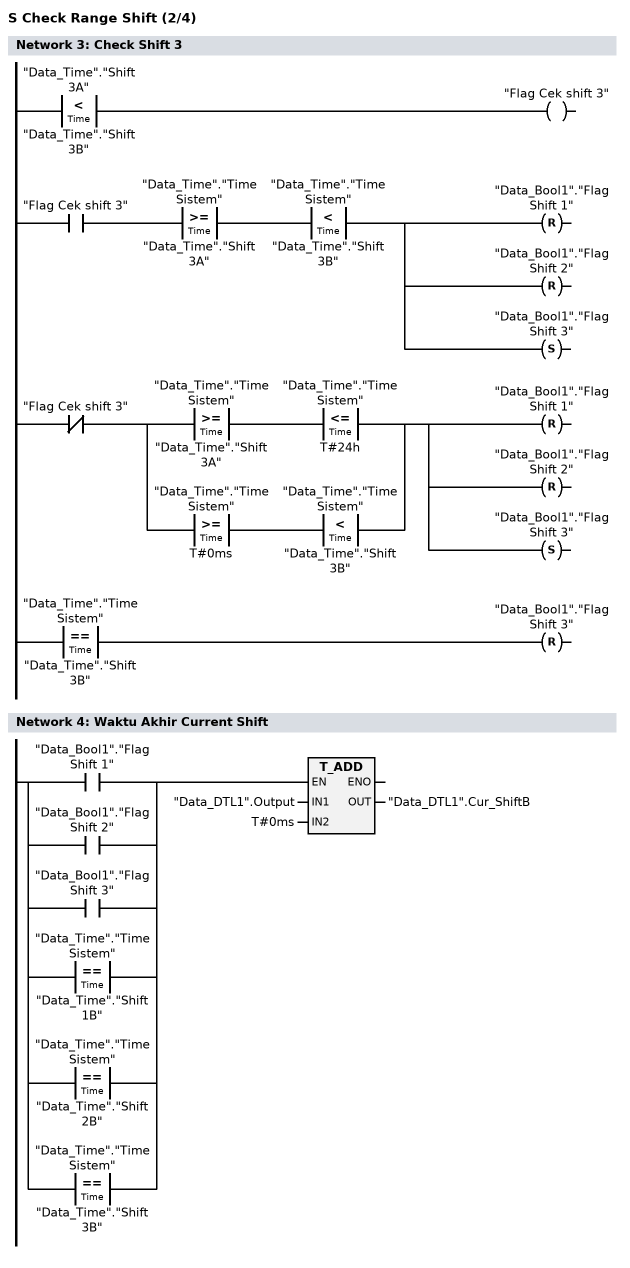
   RUNG wire#powerrail
      { S7_Templates := "SrcType := Time" } LT_Contact(in1 := "Data_Time"."Shift 3A", in2 := "Data_Time"."Shift 3B")
      Coil( "Flag Cek shift 3" )
   END_RUNG
   RUNG wire#powerrail
      Contact( "Flag Cek shift 3" )
      { S7_Templates := "SrcType := Time" } GE_Contact(in1 := "Data_Time"."Time Sistem", in2 := "Data_Time"."Shift 3A")
      { S7_Templates := "SrcType := Time" } LT_Contact(in1 := "Data_Time"."Time Sistem", in2 := "Data_Time"."Shift 3B")
      wire#w1
      R_Coil( "Data_Bool1"."Flag Shift 1" )
   END_RUNG
   RUNG wire#w1
      R_Coil( "Data_Bool1"."Flag Shift 2" )
   END_RUNG
   RUNG wire#w1
      S_Coil( "Data_Bool1"."Flag Shift 3" )
   END_RUNG
   RUNG wire#powerrail
      I_Contact( "Flag Cek shift 3" )
      wire#w2
      { S7_Templates := "SrcType := Time" } GE_Contact(in1 := "Data_Time"."Time Sistem", in2 := "Data_Time"."Shift 3A")
      { S7_Templates := "SrcType := Time" } LE_Contact(in1 := "Data_Time"."Time Sistem", in2 := T#24h)
      wire#w3
      R_Coil( "Data_Bool1"."Flag Shift 1" )
   END_RUNG
   RUNG wire#w2
      { S7_Templates := "SrcType := Time" } GE_Contact(in1 := "Data_Time"."Time Sistem", in2 := T#0ms)
      { S7_Templates := "SrcType := Time" } LT_Contact(in1 := "Data_Time"."Time Sistem", in2 := "Data_Time"."Shift 3B")
   END_RUNG wire#w3
   RUNG wire#w3
      R_Coil( "Data_Bool1"."Flag Shift 2" )
   END_RUNG
   RUNG wire#w3
      S_Coil( "Data_Bool1"."Flag Shift 3" )
   END_RUNG
   RUNG wire#powerrail
      { S7_Templates := "SrcType := Time" } EQ_Contact(in1 := "Data_Time"."Time Sistem", in2 := "Data_Time"."Shift 3B")
      R_Coil( "Data_Bool1"."Flag Shift 3" )
   END_RUNG
   // the same network as SCL:
   "Flag Cek shift 3" := "Data_Time"."Shift 3A" < "Data_Time"."Shift 3B";
   IF "Flag Cek shift 3" AND ("Data_Time"."Time Sistem" >= "Data_Time"."Shift 3A") AND ("Data_Time"."Time Sistem" < "Data_Time"."Shift 3B") THEN
       "Data_Bool1"."Flag Shift 1" := FALSE;
       "Data_Bool1"."Flag Shift 2" := FALSE;
       "Data_Bool1"."Flag Shift 3" := TRUE;
   END_IF;
   IF NOT "Flag Cek shift 3" AND ((("Data_Time"."Time Sistem" >= "Data_Time"."Shift 3A") AND ("Data_Time"."Time Sistem" <= T#24h)) OR (("Data_Time"."Time Sistem" >= T#0ms) AND ("Data_Time"."Time Sistem" < "Data_Time"."Shift 3B"))) THEN
       "Data_Bool1"."Flag Shift 1" := FALSE;
       "Data_Bool1"."Flag Shift 2" := FALSE;
       "Data_Bool1"."Flag Shift 3" := TRUE;
   END_IF;
   IF "Data_Time"."Time Sistem" = "Data_Time"."Shift 3B" THEN "Data_Bool1"."Flag Shift 3" := FALSE; END_IF;
END_REGION

REGION Network 4: Waktu Akhir Current Shift
   IF "Data_Bool1"."Flag Shift 1" OR "Data_Bool1"."Flag Shift 2" OR "Data_Bool1"."Flag Shift 3" OR ("Data_Time"."Time Sistem" = "Data_Time"."Shift 1B") OR ("Data_Time"."Time Sistem" = "Data_Time"."Shift 2B") OR ("Data_Time"."Time Sistem" = "Data_Time"."Shift 3B") THEN
       "Data_DTL1".Cur_ShiftB := T_ADD(IN1 := "Data_DTL1".Output, IN2 := T#0ms);
   END_IF;
END_REGION

REGION Network 5: Waktu Awal Current Shift
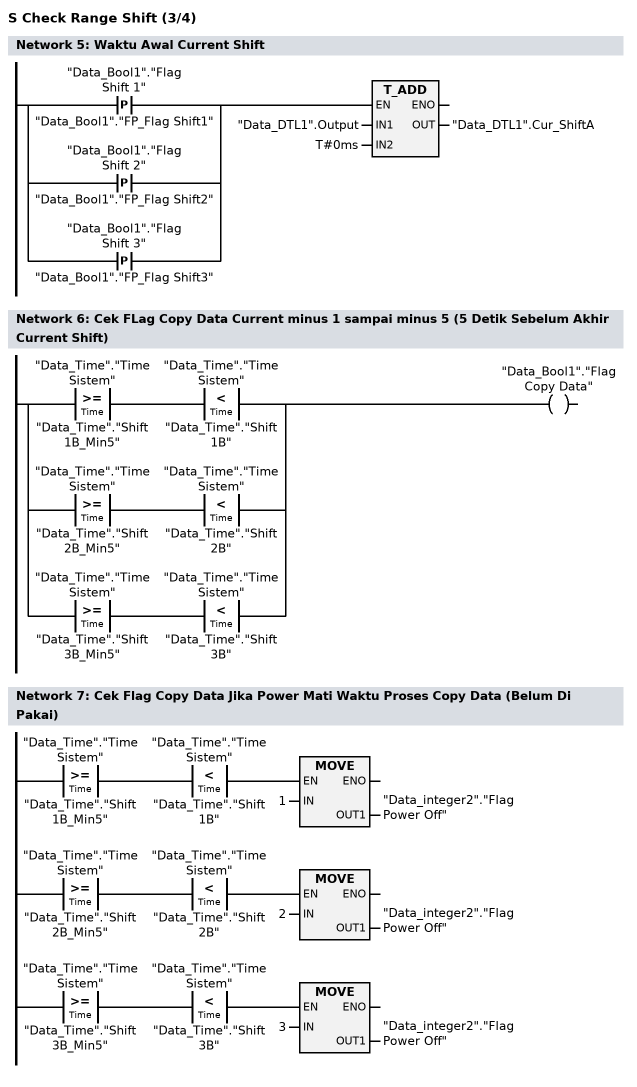
   #_w1 := "Data_Bool1"."Flag Shift 1" AND NOT "Data_Bool1"."FP_Flag Shift1";   // rising edge of "Data_Bool1"."Flag Shift 1"
   "Data_Bool1"."FP_Flag Shift1" := "Data_Bool1"."Flag Shift 1";
   #_w2 := "Data_Bool1"."Flag Shift 2" AND NOT "Data_Bool1"."FP_Flag Shift2";   // rising edge of "Data_Bool1"."Flag Shift 2"
   "Data_Bool1"."FP_Flag Shift2" := "Data_Bool1"."Flag Shift 2";
   #_w3 := "Data_Bool1"."Flag Shift 3" AND NOT "Data_Bool1"."FP_Flag Shift3";   // rising edge of "Data_Bool1"."Flag Shift 3"
   "Data_Bool1"."FP_Flag Shift3" := "Data_Bool1"."Flag Shift 3";
   IF #_w1 OR #_w2 OR #_w3 THEN
       "Data_DTL1".Cur_ShiftA := T_ADD(IN1 := "Data_DTL1".Output, IN2 := T#0ms);
   END_IF;
END_REGION

REGION Network 6: Cek FLag Copy Data Current minus 1 sampai minus 5 (5 Detik Sebelum Akhir Current Shift)
   RUNG wire#powerrail
      { S7_Templates := "SrcType := Time" } GE_Contact(in1 := "Data_Time"."Time Sistem", in2 := "Data_Time"."Shift 1B_Min5")
      { S7_Templates := "SrcType := Time" } LT_Contact(in1 := "Data_Time"."Time Sistem", in2 := "Data_Time"."Shift 1B")
      wire#w1
      Coil( "Data_Bool1"."Flag Copy Data" )
   END_RUNG
   RUNG wire#powerrail
      { S7_Templates := "SrcType := Time" } GE_Contact(in1 := "Data_Time"."Time Sistem", in2 := "Data_Time"."Shift 2B_Min5")
      { S7_Templates := "SrcType := Time" } LT_Contact(in1 := "Data_Time"."Time Sistem", in2 := "Data_Time"."Shift 2B")
   END_RUNG wire#w1
   RUNG wire#powerrail
      { S7_Templates := "SrcType := Time" } GE_Contact(in1 := "Data_Time"."Time Sistem", in2 := "Data_Time"."Shift 3B_Min5")
      { S7_Templates := "SrcType := Time" } LT_Contact(in1 := "Data_Time"."Time Sistem", in2 := "Data_Time"."Shift 3B")
   END_RUNG wire#w1
   // the same network as SCL:
   "Data_Bool1"."Flag Copy Data" := (("Data_Time"."Time Sistem" >= "Data_Time"."Shift 1B_Min5") AND ("Data_Time"."Time Sistem" < "Data_Time"."Shift 1B")) OR (("Data_Time"."Time Sistem" >= "Data_Time"."Shift 2B_Min5") AND ("Data_Time"."Time Sistem" < "Data_Time"."Shift 2B")) OR (("Data_Time"."Time Sistem" >= "Data_Time"."Shift 3B_Min5") AND ("Data_Time"."Time Sistem" < "Data_Time"."Shift 3B"));
END_REGION

REGION Network 7: Cek Flag Copy Data Jika Power Mati Waktu Proses Copy Data (Belum Di Pakai)
   RUNG wire#powerrail
      { S7_Templates := "SrcType := Time" } GE_Contact(in1 := "Data_Time"."Time Sistem", in2 := "Data_Time"."Shift 1B_Min5")
      { S7_Templates := "SrcType := Time" } LT_Contact(in1 := "Data_Time"."Time Sistem", in2 := "Data_Time"."Shift 1B")
      { S7_GenerateENO := "TRUE" } Move(in := 1, out1 => "Data_integer2"."Flag Power Off")
   END_RUNG
   RUNG wire#powerrail
      { S7_Templates := "SrcType := Time" } GE_Contact(in1 := "Data_Time"."Time Sistem", in2 := "Data_Time"."Shift 2B_Min5")
      { S7_Templates := "SrcType := Time" } LT_Contact(in1 := "Data_Time"."Time Sistem", in2 := "Data_Time"."Shift 2B")
      { S7_GenerateENO := "TRUE" } Move(in := 2, out1 => "Data_integer2"."Flag Power Off")
   END_RUNG
   RUNG wire#powerrail
      { S7_Templates := "SrcType := Time" } GE_Contact(in1 := "Data_Time"."Time Sistem", in2 := "Data_Time"."Shift 3B_Min5")
      { S7_Templates := "SrcType := Time" } LT_Contact(in1 := "Data_Time"."Time Sistem", in2 := "Data_Time"."Shift 3B")
      { S7_GenerateENO := "TRUE" } Move(in := 3, out1 => "Data_integer2"."Flag Power Off")
   END_RUNG
   // the same network as SCL:
   IF ("Data_Time"."Time Sistem" >= "Data_Time"."Shift 1B_Min5") AND ("Data_Time"."Time Sistem" < "Data_Time"."Shift 1B") THEN
       "Data_integer2"."Flag Power Off" := 1;
   END_IF;
   IF ("Data_Time"."Time Sistem" >= "Data_Time"."Shift 2B_Min5") AND ("Data_Time"."Time Sistem" < "Data_Time"."Shift 2B") THEN
       "Data_integer2"."Flag Power Off" := 2;
   END_IF;
   IF ("Data_Time"."Time Sistem" >= "Data_Time"."Shift 3B_Min5") AND ("Data_Time"."Time Sistem" < "Data_Time"."Shift 3B") THEN
       "Data_integer2"."Flag Power Off" := 3;
   END_IF;
END_REGION

REGION Network 8: Waktu Awal Current Shift Static Dan Set Copi data Setelah Power mati di waktu proses Copi Data (belum Dipakai)
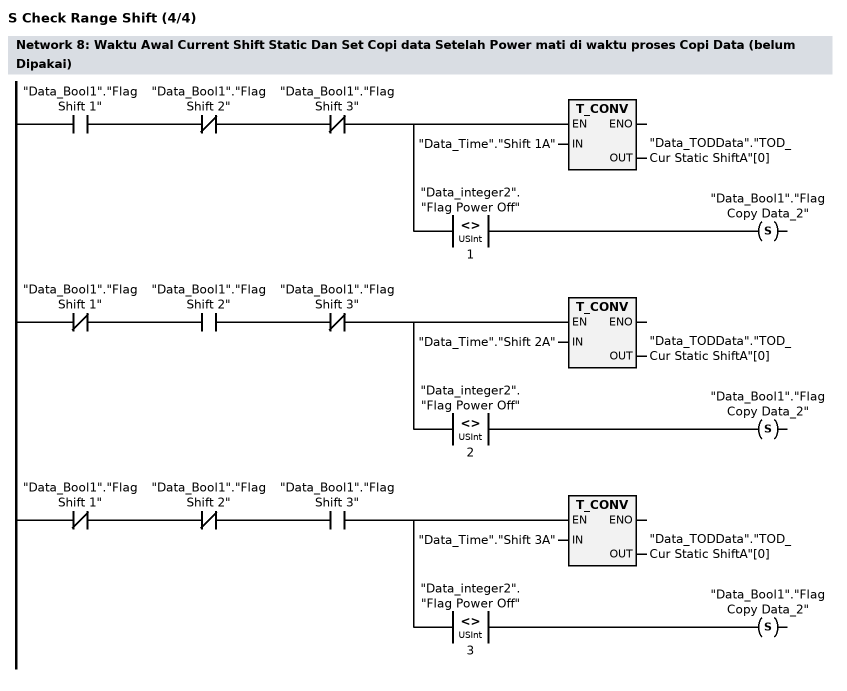
   #_w1 := "Data_Bool1"."Flag Shift 1" AND NOT "Data_Bool1"."Flag Shift 2" AND NOT "Data_Bool1"."Flag Shift 3";
   IF #_w1 THEN "Data_TODData"."TOD_Cur Static ShiftA"[0] := T_CONV(IN := "Data_Time"."Shift 1A"); END_IF;
   IF #_w1 AND ("Data_integer2"."Flag Power Off" <> 1) THEN "Data_Bool1"."Flag Copy Data_2" := TRUE; END_IF;
   #_w2 := NOT "Data_Bool1"."Flag Shift 1" AND "Data_Bool1"."Flag Shift 2" AND NOT "Data_Bool1"."Flag Shift 3";
   IF #_w2 THEN "Data_TODData"."TOD_Cur Static ShiftA"[0] := T_CONV(IN := "Data_Time"."Shift 2A"); END_IF;
   IF #_w2 AND ("Data_integer2"."Flag Power Off" <> 2) THEN "Data_Bool1"."Flag Copy Data_2" := TRUE; END_IF;
   #_w3 := NOT "Data_Bool1"."Flag Shift 1" AND NOT "Data_Bool1"."Flag Shift 2" AND "Data_Bool1"."Flag Shift 3";
   IF #_w3 THEN "Data_TODData"."TOD_Cur Static ShiftA"[0] := T_CONV(IN := "Data_Time"."Shift 3A"); END_IF;
   IF #_w3 AND ("Data_integer2"."Flag Power Off" <> 3) THEN "Data_Bool1"."Flag Copy Data_2" := TRUE; END_IF;
END_REGION
END_FUNCTION_BLOCK

FUNCTION_BLOCK "S Block Current Shift_M2"   // FB11, LAD
{ S7_Optimized_Access := 'TRUE' }
VERSION : 0.1
BEGIN

REGION Network 1: Move Data Input sloft Minus 1 To 2
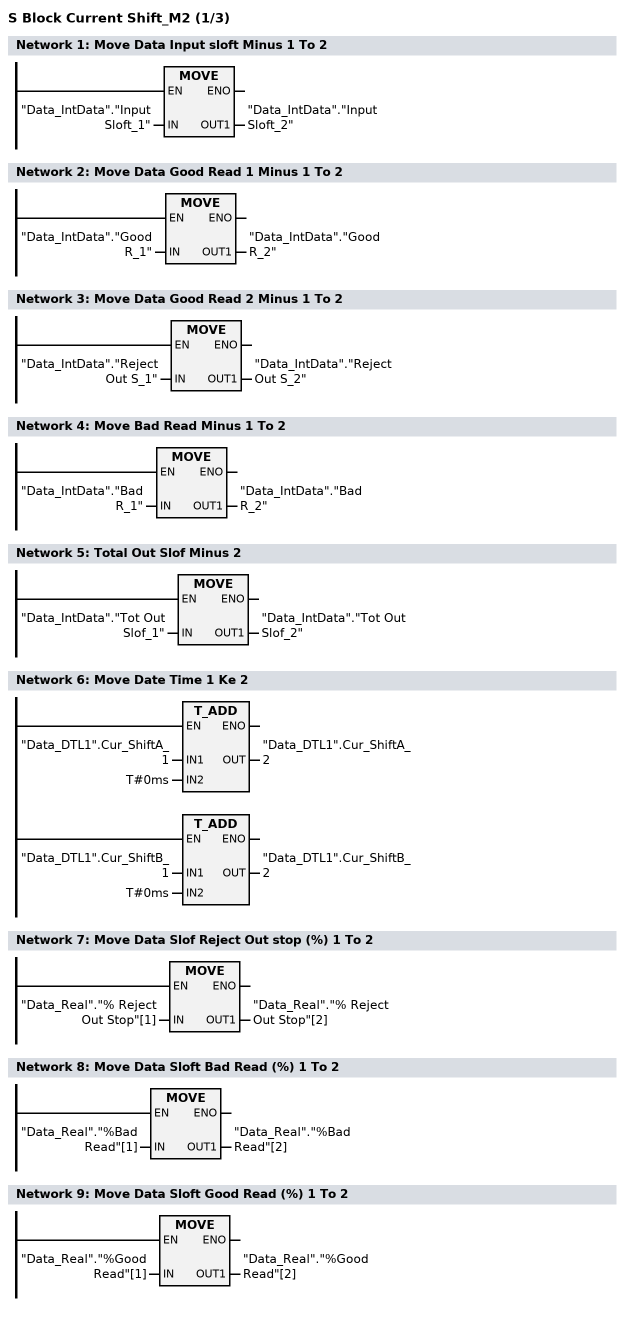
   RUNG wire#powerrail
      { S7_GenerateENO := "TRUE" } Move(in := "Data_IntData"."Input Sloft_1", out1 => "Data_IntData"."Input Sloft_2")
   END_RUNG
   // the same network as SCL:
   "Data_IntData"."Input Sloft_2" := "Data_IntData"."Input Sloft_1";
END_REGION

REGION Network 2: Move Data Good Read 1 Minus 1 To 2
   RUNG wire#powerrail
      { S7_GenerateENO := "TRUE" } Move(in := "Data_IntData"."Good R_1", out1 => "Data_IntData"."Good R_2")
   END_RUNG
   // the same network as SCL:
   "Data_IntData"."Good R_2" := "Data_IntData"."Good R_1";
END_REGION

REGION Network 3: Move Data Good Read 2 Minus 1 To 2
   RUNG wire#powerrail
      { S7_GenerateENO := "TRUE" } Move(in := "Data_IntData"."Reject Out S_1", out1 => "Data_IntData"."Reject Out S_2")
   END_RUNG
   // the same network as SCL:
   "Data_IntData"."Reject Out S_2" := "Data_IntData"."Reject Out S_1";
END_REGION

REGION Network 4: Move Bad Read Minus 1 To 2
   RUNG wire#powerrail
      { S7_GenerateENO := "TRUE" } Move(in := "Data_IntData"."Bad R_1", out1 => "Data_IntData"."Bad R_2")
   END_RUNG
   // the same network as SCL:
   "Data_IntData"."Bad R_2" := "Data_IntData"."Bad R_1";
END_REGION

REGION Network 5: Total Out Slof Minus 2
   RUNG wire#powerrail
      { S7_GenerateENO := "TRUE" } Move(in := "Data_IntData"."Tot Out Slof_1", out1 => "Data_IntData"."Tot Out Slof_2")
   END_RUNG
   // the same network as SCL:
   "Data_IntData"."Tot Out Slof_2" := "Data_IntData"."Tot Out Slof_1";
END_REGION

REGION Network 6: Move Date Time 1 Ke 2
   "Data_DTL1".Cur_ShiftA_2 := T_ADD(IN1 := "Data_DTL1".Cur_ShiftA_1, IN2 := T#0ms);
   "Data_DTL1".Cur_ShiftB_2 := T_ADD(IN1 := "Data_DTL1".Cur_ShiftB_1, IN2 := T#0ms);
END_REGION

REGION Network 7: Move Data Slof Reject Out stop (%) 1 To 2
   RUNG wire#powerrail
      { S7_GenerateENO := "TRUE" } Move(in := "Data_Real"."% Reject Out Stop"[1], out1 => "Data_Real"."% Reject Out Stop"[2])
   END_RUNG
   // the same network as SCL:
   "Data_Real"."% Reject Out Stop"[2] := "Data_Real"."% Reject Out Stop"[1];
END_REGION

REGION Network 8: Move Data Sloft Bad Read (%) 1 To 2
   RUNG wire#powerrail
      { S7_GenerateENO := "TRUE" } Move(in := "Data_Real"."%Bad Read"[1], out1 => "Data_Real"."%Bad Read"[2])
   END_RUNG
   // the same network as SCL:
   "Data_Real"."%Bad Read"[2] := "Data_Real"."%Bad Read"[1];
END_REGION

REGION Network 9: Move Data Sloft Good Read (%) 1 To 2
   RUNG wire#powerrail
      { S7_GenerateENO := "TRUE" } Move(in := "Data_Real"."%Good Read"[1], out1 => "Data_Real"."%Good Read"[2])
   END_RUNG
   // the same network as SCL:
   "Data_Real"."%Good Read"[2] := "Data_Real"."%Good Read"[1];
END_REGION

REGION Network 10: Move Output Data Total Sloft (%) 1 To 2
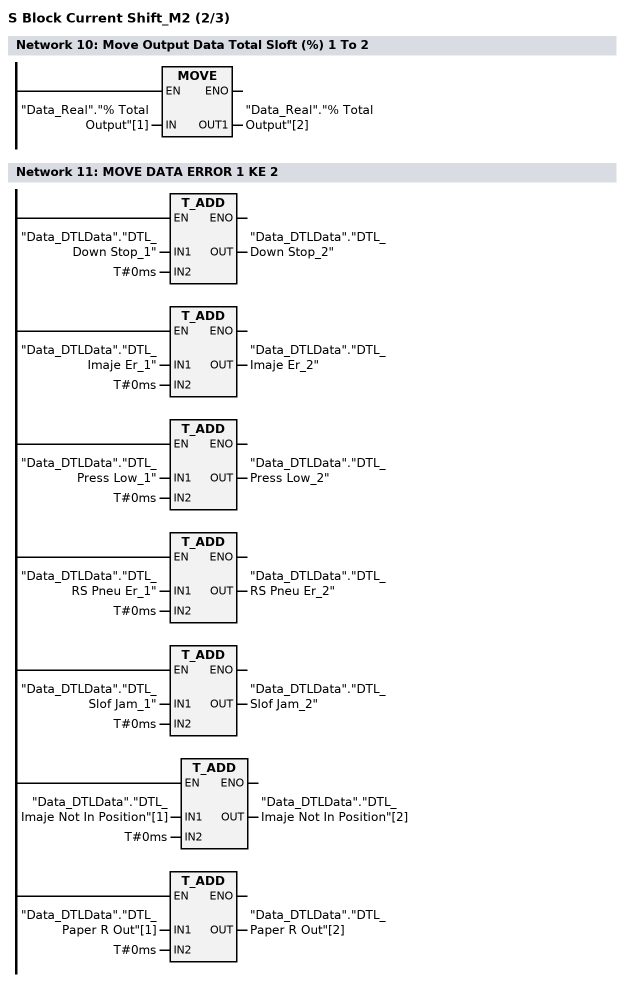
   RUNG wire#powerrail
      { S7_GenerateENO := "TRUE" } Move(in := "Data_Real"."% Total Output"[1], out1 => "Data_Real"."% Total Output"[2])
   END_RUNG
   // the same network as SCL:
   "Data_Real"."% Total Output"[2] := "Data_Real"."% Total Output"[1];
END_REGION

REGION Network 11: MOVE DATA ERROR 1 KE 2
   "Data_DTLData"."DTL_Down Stop_2" := T_ADD(IN1 := "Data_DTLData"."DTL_Down Stop_1", IN2 := T#0ms);
   "Data_DTLData"."DTL_Imaje Er_2" := T_ADD(IN1 := "Data_DTLData"."DTL_Imaje Er_1", IN2 := T#0ms);
   "Data_DTLData"."DTL_Press Low_2" := T_ADD(IN1 := "Data_DTLData"."DTL_Press Low_1", IN2 := T#0ms);
   "Data_DTLData"."DTL_RS Pneu Er_2" := T_ADD(IN1 := "Data_DTLData"."DTL_RS Pneu Er_1", IN2 := T#0ms);
   "Data_DTLData"."DTL_Slof Jam_2" := T_ADD(IN1 := "Data_DTLData"."DTL_Slof Jam_1", IN2 := T#0ms);
   "Data_DTLData"."DTL_Imaje Not In Position"[2] := T_ADD(IN1 := "Data_DTLData"."DTL_Imaje Not In Position"[1],
                           IN2 := T#0ms);
   "Data_DTLData"."DTL_Paper R Out"[2] := T_ADD(IN1 := "Data_DTLData"."DTL_Paper R Out"[1], IN2 := T#0ms);
END_REGION

REGION Network 12: Copi Data Frekuensi error
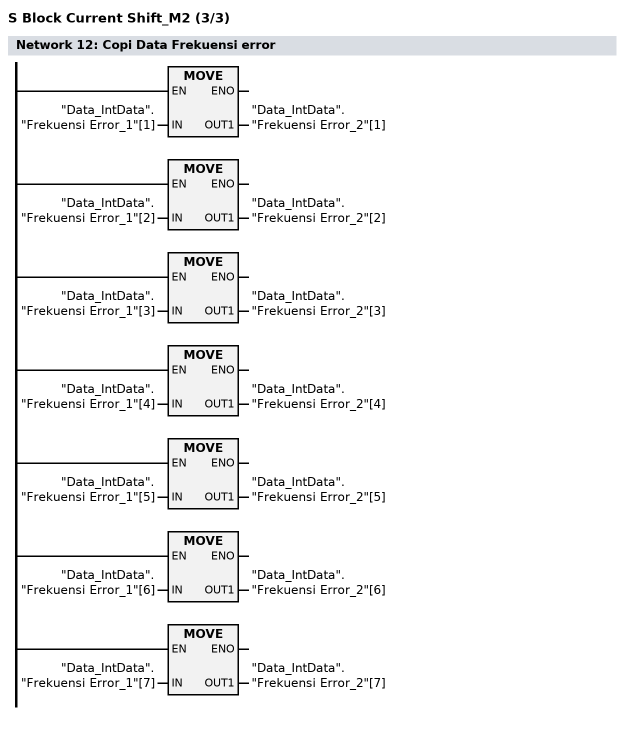
   RUNG wire#powerrail
      { S7_GenerateENO := "TRUE" } Move(in := "Data_IntData"."Frekuensi Error_1"[1], out1 => "Data_IntData"."Frekuensi Error_2"[1])
   END_RUNG
   RUNG wire#powerrail
      { S7_GenerateENO := "TRUE" } Move(in := "Data_IntData"."Frekuensi Error_1"[2], out1 => "Data_IntData"."Frekuensi Error_2"[2])
   END_RUNG
   RUNG wire#powerrail
      { S7_GenerateENO := "TRUE" } Move(in := "Data_IntData"."Frekuensi Error_1"[3], out1 => "Data_IntData"."Frekuensi Error_2"[3])
   END_RUNG
   RUNG wire#powerrail
      { S7_GenerateENO := "TRUE" } Move(in := "Data_IntData"."Frekuensi Error_1"[4], out1 => "Data_IntData"."Frekuensi Error_2"[4])
   END_RUNG
   RUNG wire#powerrail
      { S7_GenerateENO := "TRUE" } Move(in := "Data_IntData"."Frekuensi Error_1"[5], out1 => "Data_IntData"."Frekuensi Error_2"[5])
   END_RUNG
   RUNG wire#powerrail
      { S7_GenerateENO := "TRUE" } Move(in := "Data_IntData"."Frekuensi Error_1"[6], out1 => "Data_IntData"."Frekuensi Error_2"[6])
   END_RUNG
   RUNG wire#powerrail
      { S7_GenerateENO := "TRUE" } Move(in := "Data_IntData"."Frekuensi Error_1"[7], out1 => "Data_IntData"."Frekuensi Error_2"[7])
   END_RUNG
   // the same network as SCL:
   "Data_IntData"."Frekuensi Error_2"[1] := "Data_IntData"."Frekuensi Error_1"[1];
   "Data_IntData"."Frekuensi Error_2"[2] := "Data_IntData"."Frekuensi Error_1"[2];
   "Data_IntData"."Frekuensi Error_2"[3] := "Data_IntData"."Frekuensi Error_1"[3];
   "Data_IntData"."Frekuensi Error_2"[4] := "Data_IntData"."Frekuensi Error_1"[4];
   "Data_IntData"."Frekuensi Error_2"[5] := "Data_IntData"."Frekuensi Error_1"[5];
   "Data_IntData"."Frekuensi Error_2"[6] := "Data_IntData"."Frekuensi Error_1"[6];
   "Data_IntData"."Frekuensi Error_2"[7] := "Data_IntData"."Frekuensi Error_1"[7];
END_REGION
END_FUNCTION_BLOCK

FUNCTION_BLOCK "S Block Current Shift_M3"   // FB12, LAD
{ S7_Optimized_Access := 'TRUE' }
VERSION : 0.1
BEGIN

REGION Network 1: Move Data Input sloft Minus 2 To 3
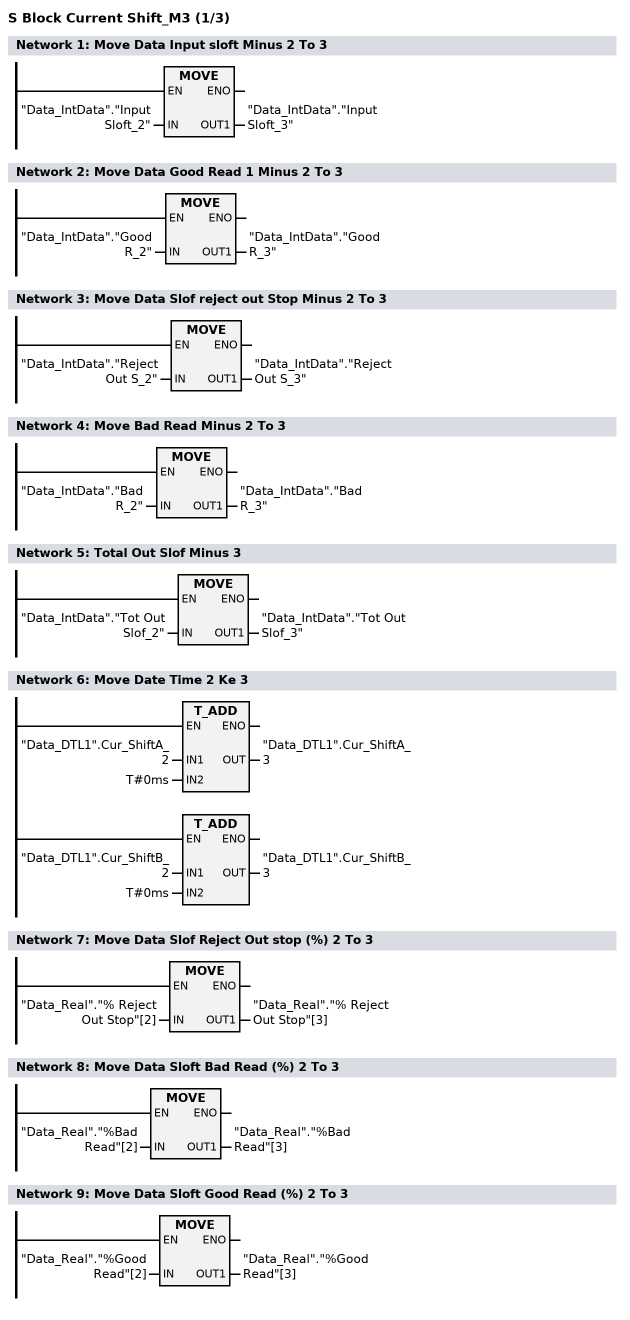
   RUNG wire#powerrail
      { S7_GenerateENO := "TRUE" } Move(in := "Data_IntData"."Input Sloft_2", out1 => "Data_IntData"."Input Sloft_3")
   END_RUNG
   // the same network as SCL:
   "Data_IntData"."Input Sloft_3" := "Data_IntData"."Input Sloft_2";
END_REGION

REGION Network 2: Move Data Good Read 1 Minus 2 To 3
   RUNG wire#powerrail
      { S7_GenerateENO := "TRUE" } Move(in := "Data_IntData"."Good R_2", out1 => "Data_IntData"."Good R_3")
   END_RUNG
   // the same network as SCL:
   "Data_IntData"."Good R_3" := "Data_IntData"."Good R_2";
END_REGION

REGION Network 3: Move Data Slof reject out Stop Minus 2 To 3
   RUNG wire#powerrail
      { S7_GenerateENO := "TRUE" } Move(in := "Data_IntData"."Reject Out S_2", out1 => "Data_IntData"."Reject Out S_3")
   END_RUNG
   // the same network as SCL:
   "Data_IntData"."Reject Out S_3" := "Data_IntData"."Reject Out S_2";
END_REGION

REGION Network 4: Move Bad Read Minus 2 To 3
   RUNG wire#powerrail
      { S7_GenerateENO := "TRUE" } Move(in := "Data_IntData"."Bad R_2", out1 => "Data_IntData"."Bad R_3")
   END_RUNG
   // the same network as SCL:
   "Data_IntData"."Bad R_3" := "Data_IntData"."Bad R_2";
END_REGION

REGION Network 5: Total Out Slof Minus 3
   RUNG wire#powerrail
      { S7_GenerateENO := "TRUE" } Move(in := "Data_IntData"."Tot Out Slof_2", out1 => "Data_IntData"."Tot Out Slof_3")
   END_RUNG
   // the same network as SCL:
   "Data_IntData"."Tot Out Slof_3" := "Data_IntData"."Tot Out Slof_2";
END_REGION

REGION Network 6: Move Date Time 2 Ke 3
   "Data_DTL1".Cur_ShiftA_3 := T_ADD(IN1 := "Data_DTL1".Cur_ShiftA_2, IN2 := T#0ms);
   "Data_DTL1".Cur_ShiftB_3 := T_ADD(IN1 := "Data_DTL1".Cur_ShiftB_2, IN2 := T#0ms);
END_REGION

REGION Network 7: Move Data Slof Reject Out stop (%) 2 To 3
   RUNG wire#powerrail
      { S7_GenerateENO := "TRUE" } Move(in := "Data_Real"."% Reject Out Stop"[2], out1 => "Data_Real"."% Reject Out Stop"[3])
   END_RUNG
   // the same network as SCL:
   "Data_Real"."% Reject Out Stop"[3] := "Data_Real"."% Reject Out Stop"[2];
END_REGION

REGION Network 8: Move Data Sloft Bad Read (%) 2 To 3
   RUNG wire#powerrail
      { S7_GenerateENO := "TRUE" } Move(in := "Data_Real"."%Bad Read"[2], out1 => "Data_Real"."%Bad Read"[3])
   END_RUNG
   // the same network as SCL:
   "Data_Real"."%Bad Read"[3] := "Data_Real"."%Bad Read"[2];
END_REGION

REGION Network 9: Move Data Sloft Good Read (%) 2 To 3
   RUNG wire#powerrail
      { S7_GenerateENO := "TRUE" } Move(in := "Data_Real"."%Good Read"[2], out1 => "Data_Real"."%Good Read"[3])
   END_RUNG
   // the same network as SCL:
   "Data_Real"."%Good Read"[3] := "Data_Real"."%Good Read"[2];
END_REGION

REGION Network 10: Move Output Data Total Sloft (%) 2 To 3
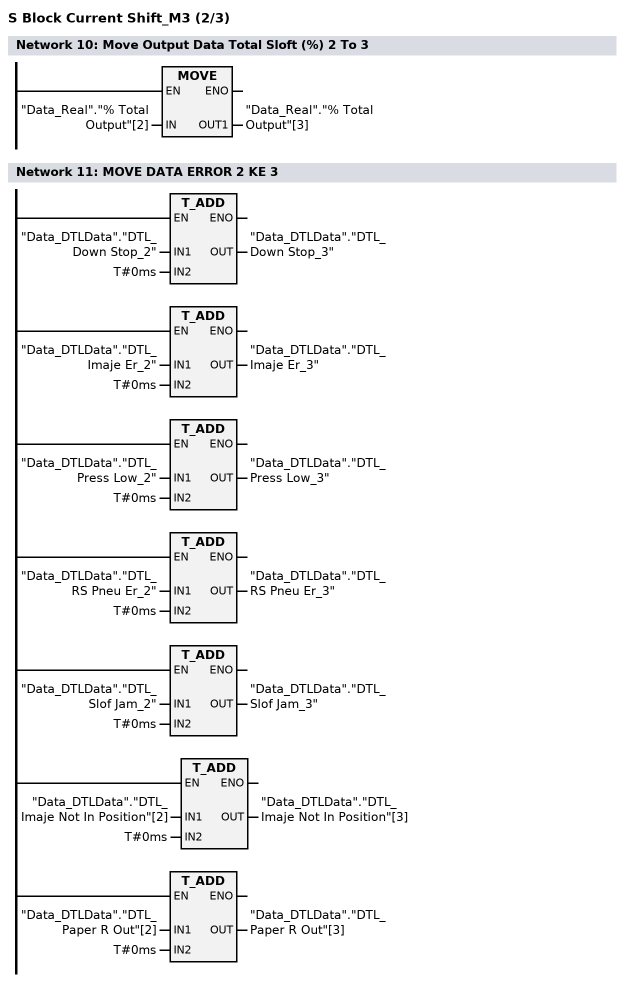
   RUNG wire#powerrail
      { S7_GenerateENO := "TRUE" } Move(in := "Data_Real"."% Total Output"[2], out1 => "Data_Real"."% Total Output"[3])
   END_RUNG
   // the same network as SCL:
   "Data_Real"."% Total Output"[3] := "Data_Real"."% Total Output"[2];
END_REGION

REGION Network 11: MOVE DATA ERROR 2 KE 3
   "Data_DTLData"."DTL_Down Stop_3" := T_ADD(IN1 := "Data_DTLData"."DTL_Down Stop_2", IN2 := T#0ms);
   "Data_DTLData"."DTL_Imaje Er_3" := T_ADD(IN1 := "Data_DTLData"."DTL_Imaje Er_2", IN2 := T#0ms);
   "Data_DTLData"."DTL_Press Low_3" := T_ADD(IN1 := "Data_DTLData"."DTL_Press Low_2", IN2 := T#0ms);
   "Data_DTLData"."DTL_RS Pneu Er_3" := T_ADD(IN1 := "Data_DTLData"."DTL_RS Pneu Er_2", IN2 := T#0ms);
   "Data_DTLData"."DTL_Slof Jam_3" := T_ADD(IN1 := "Data_DTLData"."DTL_Slof Jam_2", IN2 := T#0ms);
   "Data_DTLData"."DTL_Imaje Not In Position"[3] := T_ADD(IN1 := "Data_DTLData"."DTL_Imaje Not In Position"[2],
                           IN2 := T#0ms);
   "Data_DTLData"."DTL_Paper R Out"[3] := T_ADD(IN1 := "Data_DTLData"."DTL_Paper R Out"[2], IN2 := T#0ms);
END_REGION

REGION Network 12: Copi Data Frekuensi error
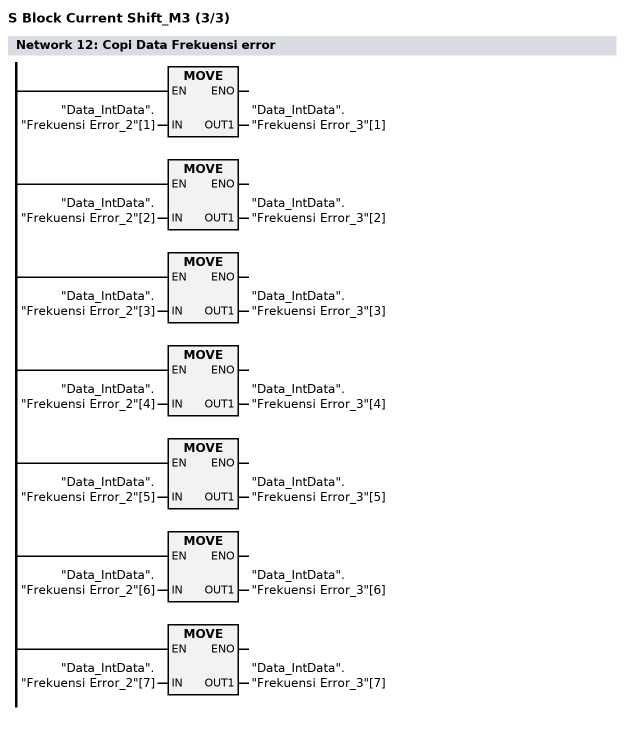
   RUNG wire#powerrail
      { S7_GenerateENO := "TRUE" } Move(in := "Data_IntData"."Frekuensi Error_2"[1], out1 => "Data_IntData"."Frekuensi Error_3"[1])
   END_RUNG
   RUNG wire#powerrail
      { S7_GenerateENO := "TRUE" } Move(in := "Data_IntData"."Frekuensi Error_2"[2], out1 => "Data_IntData"."Frekuensi Error_3"[2])
   END_RUNG
   RUNG wire#powerrail
      { S7_GenerateENO := "TRUE" } Move(in := "Data_IntData"."Frekuensi Error_2"[3], out1 => "Data_IntData"."Frekuensi Error_3"[3])
   END_RUNG
   RUNG wire#powerrail
      { S7_GenerateENO := "TRUE" } Move(in := "Data_IntData"."Frekuensi Error_2"[4], out1 => "Data_IntData"."Frekuensi Error_3"[4])
   END_RUNG
   RUNG wire#powerrail
      { S7_GenerateENO := "TRUE" } Move(in := "Data_IntData"."Frekuensi Error_2"[5], out1 => "Data_IntData"."Frekuensi Error_3"[5])
   END_RUNG
   RUNG wire#powerrail
      { S7_GenerateENO := "TRUE" } Move(in := "Data_IntData"."Frekuensi Error_2"[6], out1 => "Data_IntData"."Frekuensi Error_3"[6])
   END_RUNG
   RUNG wire#powerrail
      { S7_GenerateENO := "TRUE" } Move(in := "Data_IntData"."Frekuensi Error_2"[7], out1 => "Data_IntData"."Frekuensi Error_3"[7])
   END_RUNG
   // the same network as SCL:
   "Data_IntData"."Frekuensi Error_3"[1] := "Data_IntData"."Frekuensi Error_2"[1];
   "Data_IntData"."Frekuensi Error_3"[2] := "Data_IntData"."Frekuensi Error_2"[2];
   "Data_IntData"."Frekuensi Error_3"[3] := "Data_IntData"."Frekuensi Error_2"[3];
   "Data_IntData"."Frekuensi Error_3"[4] := "Data_IntData"."Frekuensi Error_2"[4];
   "Data_IntData"."Frekuensi Error_3"[5] := "Data_IntData"."Frekuensi Error_2"[5];
   "Data_IntData"."Frekuensi Error_3"[6] := "Data_IntData"."Frekuensi Error_2"[6];
   "Data_IntData"."Frekuensi Error_3"[7] := "Data_IntData"."Frekuensi Error_2"[7];
END_REGION
END_FUNCTION_BLOCK

FUNCTION_BLOCK "S Block Current Shift_M4"   // FB13, LAD
{ S7_Optimized_Access := 'TRUE' }
VERSION : 0.1
BEGIN

REGION Network 1: Move Data Input sloft Minus 3 To 4
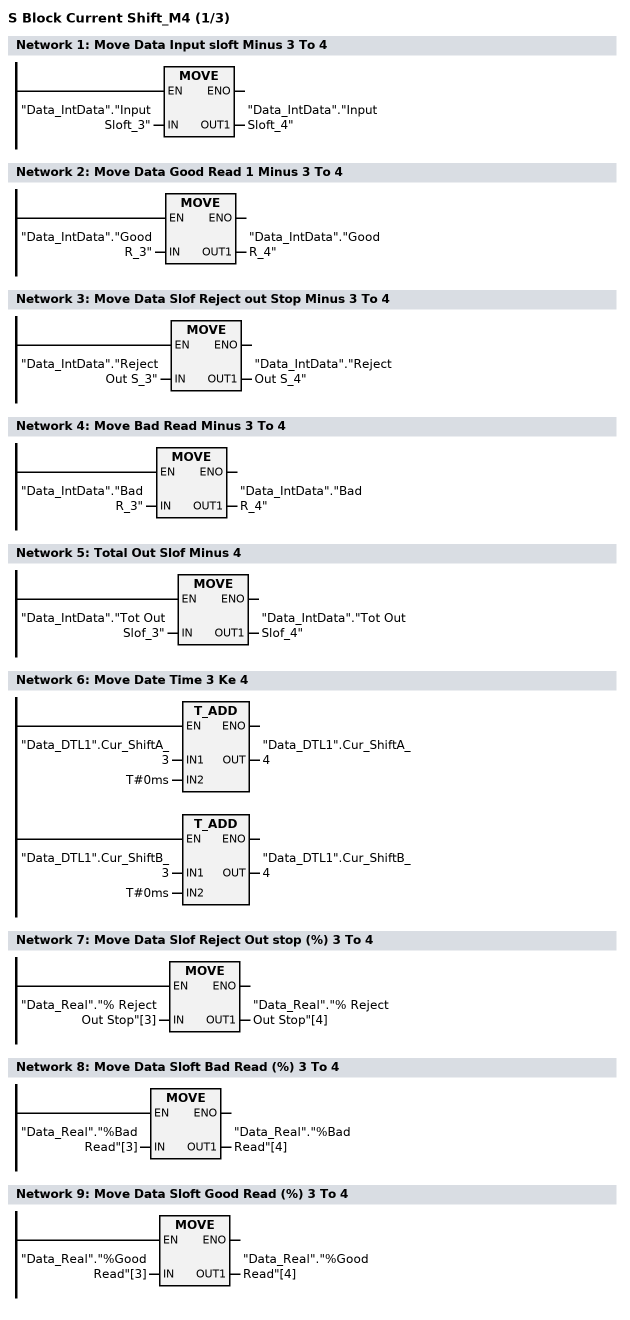
   RUNG wire#powerrail
      { S7_GenerateENO := "TRUE" } Move(in := "Data_IntData"."Input Sloft_3", out1 => "Data_IntData"."Input Sloft_4")
   END_RUNG
   // the same network as SCL:
   "Data_IntData"."Input Sloft_4" := "Data_IntData"."Input Sloft_3";
END_REGION

REGION Network 2: Move Data Good Read 1 Minus 3 To 4
   RUNG wire#powerrail
      { S7_GenerateENO := "TRUE" } Move(in := "Data_IntData"."Good R_3", out1 => "Data_IntData"."Good R_4")
   END_RUNG
   // the same network as SCL:
   "Data_IntData"."Good R_4" := "Data_IntData"."Good R_3";
END_REGION

REGION Network 3: Move Data Slof Reject out Stop Minus 3 To 4
   RUNG wire#powerrail
      { S7_GenerateENO := "TRUE" } Move(in := "Data_IntData"."Reject Out S_3", out1 => "Data_IntData"."Reject Out S_4")
   END_RUNG
   // the same network as SCL:
   "Data_IntData"."Reject Out S_4" := "Data_IntData"."Reject Out S_3";
END_REGION

REGION Network 4: Move Bad Read Minus 3 To 4
   RUNG wire#powerrail
      { S7_GenerateENO := "TRUE" } Move(in := "Data_IntData"."Bad R_3", out1 => "Data_IntData"."Bad R_4")
   END_RUNG
   // the same network as SCL:
   "Data_IntData"."Bad R_4" := "Data_IntData"."Bad R_3";
END_REGION

REGION Network 5: Total Out Slof Minus 4
   RUNG wire#powerrail
      { S7_GenerateENO := "TRUE" } Move(in := "Data_IntData"."Tot Out Slof_3", out1 => "Data_IntData"."Tot Out Slof_4")
   END_RUNG
   // the same network as SCL:
   "Data_IntData"."Tot Out Slof_4" := "Data_IntData"."Tot Out Slof_3";
END_REGION

REGION Network 6: Move Date Time 3 Ke 4
   "Data_DTL1".Cur_ShiftA_4 := T_ADD(IN1 := "Data_DTL1".Cur_ShiftA_3, IN2 := T#0ms);
   "Data_DTL1".Cur_ShiftB_4 := T_ADD(IN1 := "Data_DTL1".Cur_ShiftB_3, IN2 := T#0ms);
END_REGION

REGION Network 7: Move Data Slof Reject Out stop (%) 3 To 4
   RUNG wire#powerrail
      { S7_GenerateENO := "TRUE" } Move(in := "Data_Real"."% Reject Out Stop"[3], out1 => "Data_Real"."% Reject Out Stop"[4])
   END_RUNG
   // the same network as SCL:
   "Data_Real"."% Reject Out Stop"[4] := "Data_Real"."% Reject Out Stop"[3];
END_REGION

REGION Network 8: Move Data Sloft Bad Read (%) 3 To 4
   RUNG wire#powerrail
      { S7_GenerateENO := "TRUE" } Move(in := "Data_Real"."%Bad Read"[3], out1 => "Data_Real"."%Bad Read"[4])
   END_RUNG
   // the same network as SCL:
   "Data_Real"."%Bad Read"[4] := "Data_Real"."%Bad Read"[3];
END_REGION

REGION Network 9: Move Data Sloft Good Read (%) 3 To 4
   RUNG wire#powerrail
      { S7_GenerateENO := "TRUE" } Move(in := "Data_Real"."%Good Read"[3], out1 => "Data_Real"."%Good Read"[4])
   END_RUNG
   // the same network as SCL:
   "Data_Real"."%Good Read"[4] := "Data_Real"."%Good Read"[3];
END_REGION

REGION Network 10: Move Output Data Total Sloft (%) 3 To 4
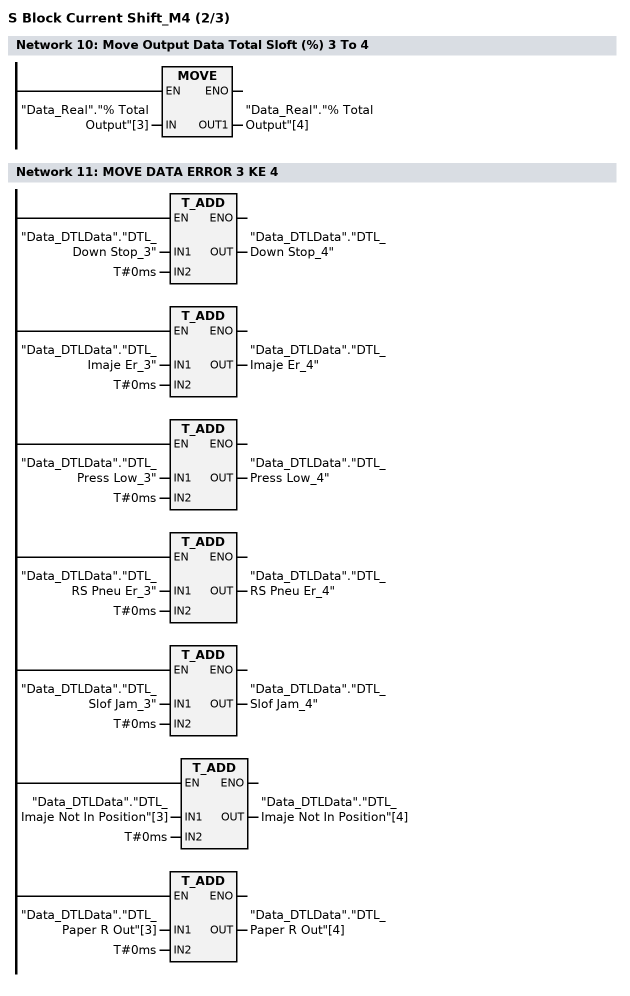
   RUNG wire#powerrail
      { S7_GenerateENO := "TRUE" } Move(in := "Data_Real"."% Total Output"[3], out1 => "Data_Real"."% Total Output"[4])
   END_RUNG
   // the same network as SCL:
   "Data_Real"."% Total Output"[4] := "Data_Real"."% Total Output"[3];
END_REGION

REGION Network 11: MOVE DATA ERROR 3 KE 4
   "Data_DTLData"."DTL_Down Stop_4" := T_ADD(IN1 := "Data_DTLData"."DTL_Down Stop_3", IN2 := T#0ms);
   "Data_DTLData"."DTL_Imaje Er_4" := T_ADD(IN1 := "Data_DTLData"."DTL_Imaje Er_3", IN2 := T#0ms);
   "Data_DTLData"."DTL_Press Low_4" := T_ADD(IN1 := "Data_DTLData"."DTL_Press Low_3", IN2 := T#0ms);
   "Data_DTLData"."DTL_RS Pneu Er_4" := T_ADD(IN1 := "Data_DTLData"."DTL_RS Pneu Er_3", IN2 := T#0ms);
   "Data_DTLData"."DTL_Slof Jam_4" := T_ADD(IN1 := "Data_DTLData"."DTL_Slof Jam_3", IN2 := T#0ms);
   "Data_DTLData"."DTL_Imaje Not In Position"[4] := T_ADD(IN1 := "Data_DTLData"."DTL_Imaje Not In Position"[3],
                           IN2 := T#0ms);
   "Data_DTLData"."DTL_Paper R Out"[4] := T_ADD(IN1 := "Data_DTLData"."DTL_Paper R Out"[3], IN2 := T#0ms);
END_REGION

REGION Network 12: Copi Data Frekuensi Error
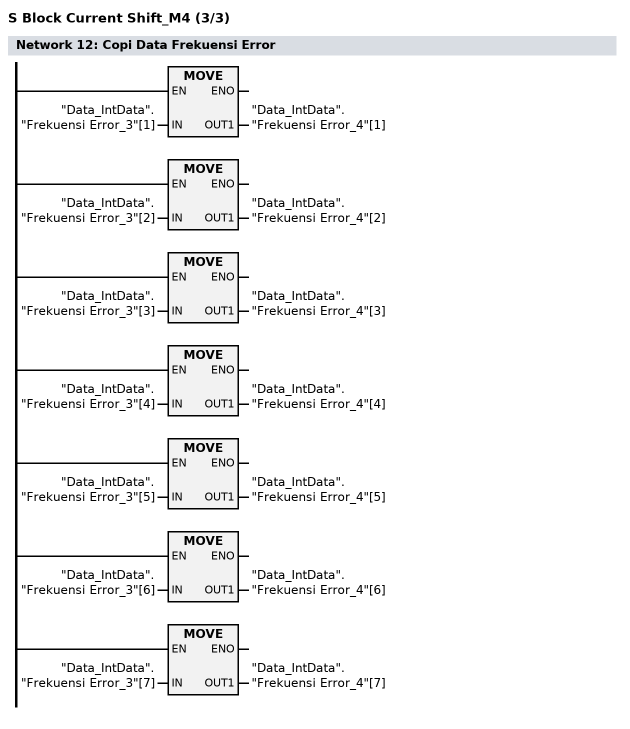
   RUNG wire#powerrail
      { S7_GenerateENO := "TRUE" } Move(in := "Data_IntData"."Frekuensi Error_3"[1], out1 => "Data_IntData"."Frekuensi Error_4"[1])
   END_RUNG
   RUNG wire#powerrail
      { S7_GenerateENO := "TRUE" } Move(in := "Data_IntData"."Frekuensi Error_3"[2], out1 => "Data_IntData"."Frekuensi Error_4"[2])
   END_RUNG
   RUNG wire#powerrail
      { S7_GenerateENO := "TRUE" } Move(in := "Data_IntData"."Frekuensi Error_3"[3], out1 => "Data_IntData"."Frekuensi Error_4"[3])
   END_RUNG
   RUNG wire#powerrail
      { S7_GenerateENO := "TRUE" } Move(in := "Data_IntData"."Frekuensi Error_3"[4], out1 => "Data_IntData"."Frekuensi Error_4"[4])
   END_RUNG
   RUNG wire#powerrail
      { S7_GenerateENO := "TRUE" } Move(in := "Data_IntData"."Frekuensi Error_3"[5], out1 => "Data_IntData"."Frekuensi Error_4"[5])
   END_RUNG
   RUNG wire#powerrail
      { S7_GenerateENO := "TRUE" } Move(in := "Data_IntData"."Frekuensi Error_3"[6], out1 => "Data_IntData"."Frekuensi Error_4"[6])
   END_RUNG
   RUNG wire#powerrail
      { S7_GenerateENO := "TRUE" } Move(in := "Data_IntData"."Frekuensi Error_3"[7], out1 => "Data_IntData"."Frekuensi Error_4"[7])
   END_RUNG
   // the same network as SCL:
   "Data_IntData"."Frekuensi Error_4"[1] := "Data_IntData"."Frekuensi Error_3"[1];
   "Data_IntData"."Frekuensi Error_4"[2] := "Data_IntData"."Frekuensi Error_3"[2];
   "Data_IntData"."Frekuensi Error_4"[3] := "Data_IntData"."Frekuensi Error_3"[3];
   "Data_IntData"."Frekuensi Error_4"[4] := "Data_IntData"."Frekuensi Error_3"[4];
   "Data_IntData"."Frekuensi Error_4"[5] := "Data_IntData"."Frekuensi Error_3"[5];
   "Data_IntData"."Frekuensi Error_4"[6] := "Data_IntData"."Frekuensi Error_3"[6];
   "Data_IntData"."Frekuensi Error_4"[7] := "Data_IntData"."Frekuensi Error_3"[7];
END_REGION
END_FUNCTION_BLOCK

FUNCTION_BLOCK "S Block Current Shift_M5"   // FB14, LAD
{ S7_Optimized_Access := 'TRUE' }
VERSION : 0.1
BEGIN

REGION Network 1: Move Data Input sloft Minus 4 To 5
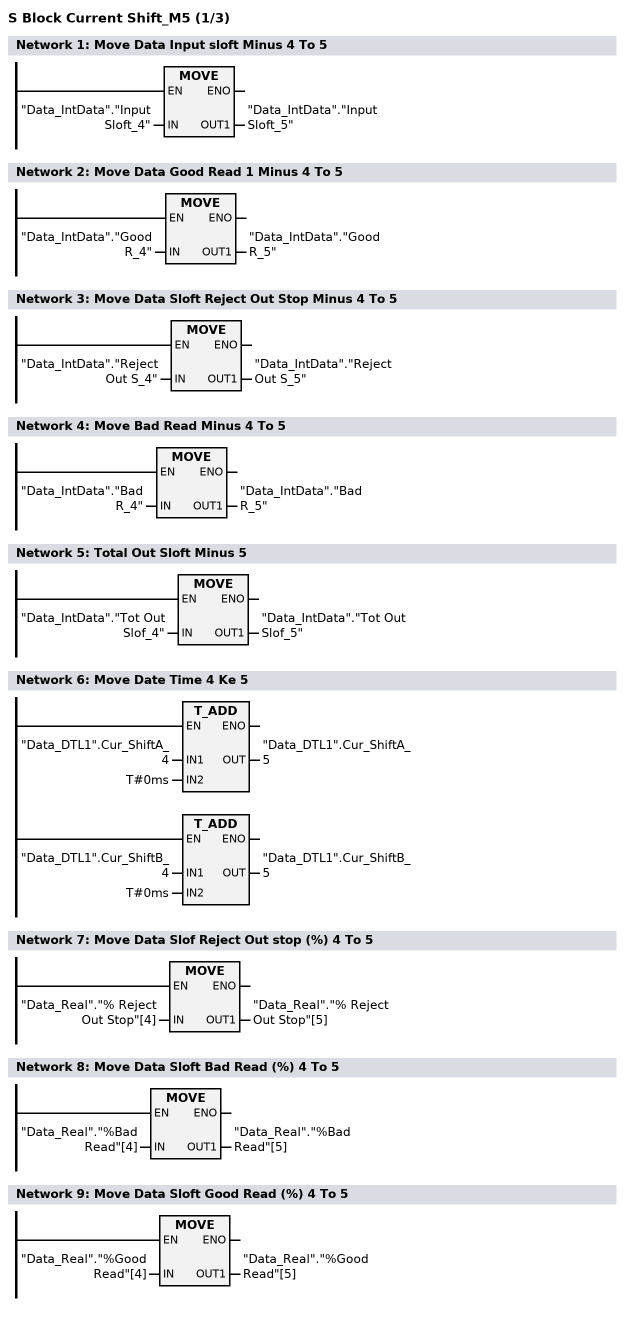
   RUNG wire#powerrail
      { S7_GenerateENO := "TRUE" } Move(in := "Data_IntData"."Input Sloft_4", out1 => "Data_IntData"."Input Sloft_5")
   END_RUNG
   // the same network as SCL:
   "Data_IntData"."Input Sloft_5" := "Data_IntData"."Input Sloft_4";
END_REGION

REGION Network 2: Move Data Good Read 1 Minus 4 To 5
   RUNG wire#powerrail
      { S7_GenerateENO := "TRUE" } Move(in := "Data_IntData"."Good R_4", out1 => "Data_IntData"."Good R_5")
   END_RUNG
   // the same network as SCL:
   "Data_IntData"."Good R_5" := "Data_IntData"."Good R_4";
END_REGION

REGION Network 3: Move Data Sloft Reject Out Stop Minus 4 To 5
   RUNG wire#powerrail
      { S7_GenerateENO := "TRUE" } Move(in := "Data_IntData"."Reject Out S_4", out1 => "Data_IntData"."Reject Out S_5")
   END_RUNG
   // the same network as SCL:
   "Data_IntData"."Reject Out S_5" := "Data_IntData"."Reject Out S_4";
END_REGION

REGION Network 4: Move Bad Read Minus 4 To 5
   RUNG wire#powerrail
      { S7_GenerateENO := "TRUE" } Move(in := "Data_IntData"."Bad R_4", out1 => "Data_IntData"."Bad R_5")
   END_RUNG
   // the same network as SCL:
   "Data_IntData"."Bad R_5" := "Data_IntData"."Bad R_4";
END_REGION

REGION Network 5: Total Out Sloft Minus 5
   RUNG wire#powerrail
      { S7_GenerateENO := "TRUE" } Move(in := "Data_IntData"."Tot Out Slof_4", out1 => "Data_IntData"."Tot Out Slof_5")
   END_RUNG
   // the same network as SCL:
   "Data_IntData"."Tot Out Slof_5" := "Data_IntData"."Tot Out Slof_4";
END_REGION

REGION Network 6: Move Date Time 4 Ke 5
   "Data_DTL1".Cur_ShiftA_5 := T_ADD(IN1 := "Data_DTL1".Cur_ShiftA_4, IN2 := T#0ms);
   "Data_DTL1".Cur_ShiftB_5 := T_ADD(IN1 := "Data_DTL1".Cur_ShiftB_4, IN2 := T#0ms);
END_REGION

REGION Network 7: Move Data Slof Reject Out stop (%) 4 To 5
   RUNG wire#powerrail
      { S7_GenerateENO := "TRUE" } Move(in := "Data_Real"."% Reject Out Stop"[4], out1 => "Data_Real"."% Reject Out Stop"[5])
   END_RUNG
   // the same network as SCL:
   "Data_Real"."% Reject Out Stop"[5] := "Data_Real"."% Reject Out Stop"[4];
END_REGION

REGION Network 8: Move Data Sloft Bad Read (%) 4 To 5
   RUNG wire#powerrail
      { S7_GenerateENO := "TRUE" } Move(in := "Data_Real"."%Bad Read"[4], out1 => "Data_Real"."%Bad Read"[5])
   END_RUNG
   // the same network as SCL:
   "Data_Real"."%Bad Read"[5] := "Data_Real"."%Bad Read"[4];
END_REGION

REGION Network 9: Move Data Sloft Good Read (%) 4 To 5
   RUNG wire#powerrail
      { S7_GenerateENO := "TRUE" } Move(in := "Data_Real"."%Good Read"[4], out1 => "Data_Real"."%Good Read"[5])
   END_RUNG
   // the same network as SCL:
   "Data_Real"."%Good Read"[5] := "Data_Real"."%Good Read"[4];
END_REGION

REGION Network 10: Move Output Data Total Sloft (%) 4 To 5
